TYPE "UDT_ZoneStructure"
VERSION : 0.1
   STRUCT
      SpeedZoneStart : DWord;
      SpeedZoneEnd : DWord;
      Zone : Word;
      Description : String[10];
      LastZone : Bool;
      StartPos : DWord;
      SpeedZone : Bool;
      NextZone : Int;
      PrevZone : Int;
      EndPos : DWord;
      AccumZone : Bool;
      ProductionZone : Bool;
      ProductionZoneSpacing : Word;
      MaxCarriers : Word;
      CarrierSpacing : Word;
      ClearToEnter : Bool;
      ClearOfStop : Bool;
      ClearZoneStart : Bool;
      ZoneFull : Bool;
      CarrierZnStatus : Array[0..60] of "UDT_ZoneCarrierStatus";
      CarrierZnStatusUnsorted : Array[0..60] of "UDT_ZoneCarrierStatus";
      InPositionTolerance : Word;
      NextCarrierClrHighSpeed : Word;
      DecelPositionOffset : Word;
      GapSpacingFault : Bool;
      GapFaultZnPosition : Int;
      GapFaultInZone : Int;
      FirstCarrierNumGapFlt : Int;
      SecondCarrierNumGapFlt : Int;
      FinePosStopZone : Bool;
      FineInPosTolerance : Word;
      FinePositionDecelOffset : Word;
      CoarseInPosTolerance : Word;
      CoarsePositionDecelOffset : Word;
      ZoneLength : Word;
      HMIZonePositionStatus : Array[1..20] of "UDT_HMIZonePositionStructure";
      HMIZonePositions : Array[1..20] of "UDT_HMIZonePositions";
      CarrierAtStop : Bool;
      CarrierNumAtStop : Word;
      StopControlFromEMS01 : "UDT_StopControlFromEMS01";
      ClearOfStopPos : DWord;
      StopStatusToEMS01 : "UDT_StopStatusToEMS01";
   END_STRUCT;
END_TYPE

TYPE "UDT_CarrierStructure"
VERSION : 0.1
   STRUCT
      SDC_IN : "UDT_SDC_IN";
      SDC_OUT : "UDT_SDC_OUT";
      ZoneFound : Word;
      Position : DWord;
      SpeedSelect : Word;
      MoveFWD : Bool;
      InProductionHold : Bool;
      Zone : Word;
      Area : String[2];
      AutoSpeedFast : Word;
      AutoSpeedSlow : Word;
      InPositionTolerance : Word;
      DecelSpeed : Word;
      DecelStartPos : DWord;
      ZonePosition : Word;
      CommFlt : Bool;
      CarrierPosition : DWord;
      CarrierNumber : Word;
      FaultsMasked : Bool;
      Faulted : Bool;
   END_STRUCT;
END_TYPE

TYPE "UDT_Zone"
VERSION : 0.1
   STRUCT
      ZONE : Array[1..60] of "UDT_ZoneStructure";
   END_STRUCT;
END_TYPE

TYPE "UDT_ZoneCarrierStatus"
VERSION : 0.1
   STRUCT
      CarrierNumber : Word;
      Position : DWord;
      RunningFWD : Bool;
   END_STRUCT;
END_TYPE

TYPE "UDT_OUT"
   STRUCT
      DecrementCarrierIndex : Bool;
      IncrementCarrierIndex : Bool;
      CarrierStatusIndex : Int;
      DecrementStatusIndex : Bool;
      IncrementStatusIndex : Bool;
      DriveStatusIndex : Int;
      DecrementZoneIndex : Bool;
      IncrementZoneIndex : Bool;
      ZoneStatusIndex : Int;
   END_STRUCT;
END_TYPE

TYPE "UDT_Carrier_Drive_Data"
   STRUCT
      CARRIER : Array[1..99] of "UDT_Drive_Data";
   END_STRUCT;
END_TYPE

TYPE "UDT_Drive_Data"
   STRUCT
      Drive_Control : Word;
      Drive_Status : Word;
   END_STRUCT;
END_TYPE

TYPE "UDT_Carrier_IO_HMI"
   STRUCT
      Carrier_Slot02_Inputs : Byte;
      Carrier_Slot03_Outputs : Byte;
      Carrier_Slot04_Inputs : Word;
      Carrier_Slot05_Outputs : Word;
   END_STRUCT;
END_TYPE

TYPE "UDT_IO_Data"
   STRUCT
      Slot2SafeInputs : Byte;
      Slot3SafeOutputs : Byte;
      Slot4StdInputs : Word;
      Slot5StdOutputs : Word;
   END_STRUCT;
END_TYPE

TYPE "UDT_Carrier_IO_Data"
   STRUCT
      CARRIER : Array[1..99] of "UDT_IO_Data";
   END_STRUCT;
END_TYPE

TYPE "UDT_Carrier_Status_HMI"
   STRUCT
      CarrierPosition : DWord;
      ActualSpeed : Word;
      RunningFWD : Bool;
      RunningREV : Bool;
      ProductionHoldPB_Status : Bool;
      CrashDetectStatus : Bool;
      AutoMode : Bool;
      ManualMode : Bool;
      DriveFwdCMD : Bool;
      DriveCmdSpeed : Word;
      NextCarrierNum : Word;
      NextStopPosition : DWord;
      Zone : Int;
      Area : String[2];
      CarrierFaultCode : Int;
      AtCmdPos : Bool;
      CommFlt : Bool;
      Faulted : Bool;
      CarrierStatusIndex : Int;
      DriveStatusIndex : Int;
      ZoneStatusIndex : Int;
      EncoderCommFault : Bool;
      DriveCommFault : Bool;
      HMICommFault : Bool;
      SetMaskCarrierFaultsPB : Bool;
      MaskCarrierFaultsLT : Bool;
      ResetMaskCarrierFaultsPB : Bool;
   END_STRUCT;
END_TYPE

TYPE "UDT_Zone_Status_HMI"
   STRUCT
      ZoneIndex : Int;
      ZoneType : String;
      NextZoneNumber : Int;
      ZoneStartPosition : DWord;
      ZoneEndPosition : DWord;
      ZoneFull : Bool;
      SpeedZone : Bool;
      SpeedZoneStartPos : DWord;
      SpeedZoneEndPos : DWord;
      AccumZoneSpacing : Word;
      ProductionZoneSpacing : Word;
      CarrierZoneStatus : Array[0..60] of "UDT_ZoneCarrierStatus";
   END_STRUCT;
END_TYPE

TYPE "UDT_StopStatusToEMS01"
   STRUCT
      StopOpen : Bool;
      StopClosed : Bool;
      CarrierAtStop : Bool;
      CarrierReleasingFromStop : Bool;
   END_STRUCT;
END_TYPE

TYPE "UDT_StopControlFromEMS01"
   STRUCT
      ClearToOpen : Bool;
      ClearToReleaseCarrier : Bool;
   END_STRUCT;
END_TYPE

TYPE "UDT_G120D_STW1_CONTROL"
VERSION : 0.1
   STRUCT
      Bit_08_JOG_R : Bool;   // 1=tippen rechtsseitig EIN/ 0= AUS / 1=jogging on right-hand side ON/ 0= OFF
      Bit_09_JOG_L : Bool;   // 1=tippen linksseitig EIN/ 0= AUS / 1=jogging on left-hand side ON/ 0= OFF
      Bit_10_CONTR_PLC : Bool;   // 1=Bedienung über PLC erforderlich/ 0=keine Bedienung über PLC erforderlich / 1=control by PLC required/ 0=no control by PLC required
      Bit_11_REVERSE : Bool;   // 1=Umkehrung des Sollwerts/ 0=keine Umkehrung / 1=inversion of setpoint/ 0=no inversion of setpoint
      Bit_12_BRAKE_Release : Bool;   // 1= Löse Bremse / 1= Release Break / 1= Manual Brake Release
      Bit_13_DDS : Bool;   // 1=DDS1 FU Datenset / 0=DDS0 FU Datenset / 1=DDS1 FU Dataset / 0=DDS0 FU Dataset
      Bit_14_DO0 : Bool;   // 1=Digitaler Ausgang aktiv/ 0=Digitaler Ausgang nicht aktiv / 1=Digital Output activ/ 0=Digital Output not activ
      Bit_15_DO1 : Bool;   // 1=Digitaler Ausgang aktiv/ 0=Digitaler Ausgang nicht aktiv / 1=Digital Output activ/ 0=Digital Output not activ
      Bit_00_ON : Bool;   // 1=EIN/ 0=AUS / 1=ON/ 0=OFF2
      Bit_01_AUS2_INH : Bool;   // 1=Betriebsvoraussetzung/ 0=AUS2 - Pulsverzögerer, Spannung auf einmal aus / 1=operation condition/ 0=AUS2 - pulse inhibitor, voltage off at once
      Bit_02_AUS3_STOP : Bool;   // 1=Betriebsvoraussetzung / 0=AUS3 - schneller Halt / 1=operation condition / 0=AUS3 - fast stop
      Bit_03_EN : Bool;   // 1=Freigabe Betrieb/ 0=deaktiviere Betrieb / 1=enable operation/ 0=disable operation
      Bit_04_EN_RAMP : Bool;   // 1=1=Betriebsvoraussetzung / 0=deaktiviere Funktionsrampengenerator / 1=operation condition / 0=disable ramp function generator
      Bit_05_START_RAMP : Bool;   // 1=Aktiviere Rampenfunktion / 0=deaktivere RFG / 1=enable ramp function generator / 0=stoppen RFG
      Bit_06_SETPOINT : Bool;   // 1=Freigabe Sollwert/ 0=deaktiviere Sollwert / 1=enable setpoint/ 0=disable setpoint
      Bit_07_RESET : Bool;   // 1=Störung quittieren / 0= irrelevant / 1=Reset fault / 0= irrelevant
   END_STRUCT;
END_TYPE

TYPE "UDT_G120D_ZSW1_STATUS"
VERSION : 0.1
   STRUCT
      Bit_08_NO_DEVIATION : Bool;   // 1=keine Abweichung des Sollwerts / 0=Abweichung / 1=no deviation current-setpoint / 0=deviation / Setpoint / actual value deviation within the tolerance range.
      Bit_09_CONTR_PLC : Bool;   // 1=Kontrolle über PLC erforderlich/ 0=keine Kontrolle erforderlich / 1=control by PLC required/ 0=no control by PLC required / The automation system is requested to ac-cept the inverter control.
      Bit_10_F_MAX : Bool;   // 1=fmax erreicht/ 0= unter fmax / 1=fmax reached/ 0= below fmax / Speed is greater than or equal to the corre-sponding maximum speed.
      Bit_11_LIMIT_REACHED : Bool;   // 1=keine Warnung/ 0=Warnung: Motor an Spannungsgrenze / 1=no warning/ 0=warning:Motor at limit of current / Comparison value for current or torque has been reached or exceeded.
      Bit_12_BRAKE_OPEN : Bool;   // 1= / 0=Haltebremse / motor Brake is open
      Bit_13_NO_OVERTEMP : Bool;   // 1= / 0=Motorüberlast / Drive Overtemperature
      Bit_14_CW_CCW : Bool;   // 1=Rechtslauf/ 0=Linkslauf / On for drive runnin clockwise/off counterclockwise
      Bit_15_OVERL : Bool;   // 1= /0= Konvertierer Überlast / 1= /0= Konverter overload / 0 = Alarm, in-verter thermal overload/on CDS display
      Bit_00_READY_RUN : Bool;   // 1=bereit zum betreiben/ 0= nicht bereit / 1=ready to run/ 0= not ready to run / Power supply switched on; electronics initial-ized; pulses locked.
      Bit_01_READY_ON : Bool;   // 1=bereit zum einschalten/ 0= nicht bereit / 1=ready to switch on/ 0= not ready to switch on / Motor is switched on (ON/OFF1 = 1), no fault is active. With the command "Enable opera-tion" (STW1.3), the inverter switches on the motor.
      Bit_02_ENABLE : Bool;   // 1=Freigabe Bedienung / 0=deaktiviere Bedienung / 1=operation enabled / 0=operation disabled / Motor follows setpoint. See control word 1, bit 3.
      Bit_03_FAULT : Bool;   // 1=Störung / 0=keine Störung / 1=fault / 0=no fault / The inverter has a fault. Acknowledge fault using STW1.7
      Bit_04_OFF2 : Bool;   // 1=kein AUS2 / 0=AUS2 Befehl ist vorhanden / 1=no AUS2 / 0=AUS2 command is present / OFF2 Coast down to standstill is not active.
      Bit_05_OFF3 : Bool;   // 1=kein AUS3 / 0=AUS3 Befehl ist vorhanden / 1=no AUS3 / 0=AUS3 command is present / OFF3 Quick stop is not active.
      Bit_06_LOCK_OUT : Bool;   // 1=sperre Ausschaltung / 0=keine Sperrung / 1=closing lock-out / 0=no closing lock-out / It is only possible to switch on the motor after an OFF1 followed by ON.
      Bit_07_WARN : Bool;   // 1=Warnung / 0= keine Warnung / 1=Warning / 0= no warning
   END_STRUCT;
END_TYPE

TYPE "UDT_G120D_ERRORS"
VERSION : 0.1
   STRUCT
      F_X33_F1 : Bool;   // Fehler Überstrom
      F_X34_F2 : Bool;   // Fehler Überspannung
      F_X35_F3 : Bool;   // Fehler Unterspannung
      F_X36_F4 : Bool;   // Fehler Inverter Übertemperatur
      F_X37_F41 : Bool;   // Fehler Motordatenerkennung
      F_X38_F52 : Bool;   // Fehler Leistungsteil
      F_X39_F62 : Bool;   // Fehler MMC Daten sind fehlerhaft
      F_X40_F70 : Bool;   // Fehler PLC Sollposition
      F_X41_F71 : Bool;   // Fehler USS Sollposition, Überwachung
      F_X42_F72 : Bool;   // Fehler USS Sollposition, USS Master
      F_X43_F90 : Bool;   // Fehler Gebersignal
      F_X44_F395 : Bool;   // Fehler CU/PM wechsel
      bit_14 : Bool;   // Reserve
      bit_15 : Bool;   // Reserve
      bit_16 : Bool;   // Reserve
      bit_17 : Bool;   // Reserve
   END_STRUCT;
END_TYPE

TYPE "UDT_SDC_EMS_FLAGS"
VERSION : 0.1
   STRUCT
      PRESENT : Bool;   // EMS vorhanden
      IN_HW : Bool;   // EMS in HardwareConfiguration
      ACTIV : Bool;   // EMS activiert
      ENABLE : Bool;   // EMS enable
      COMM_FAULT : Bool;   // EMS communicationsfehler
      FAULTY : Bool;   // EMS fehlerhaft
      SIMULATION : Bool;   // EMS simualtion
      Spare_0_7 : Bool;   // Spare
      Spare_1_0 : Bool;   // Spare
      Spare_1_1 : Bool;   // Spare
      Spare_1_2 : Bool;   // Spare
      Spare_1_3 : Bool;   // Spare
      Spare_1_4 : Bool;   // Spare
      Spare_1_5 : Bool;   // Spare
      Spare_1_6 : Bool;   // Spare
      Spare_1_7 : Bool;   // Spare
   END_STRUCT;
END_TYPE

TYPE "UDT_SDC_TS_PARAMETER"
VERSION : 0.1
   STRUCT
      ALLG : "UDT_SDC_TS_PAR_ALLG";   // allgemeine Sections Parameter
      PROFIL : Array[1..10] of "UDT_SDC_TS_PAR_PROFIL";   // Profilbezogene Sections Parameter
   END_STRUCT;
END_TYPE

TYPE "UDT_SDC_TS_PAR_PROFIL"
VERSION : 0.1
   STRUCT
      Hoist_Pos_start : Int;   // Start of hoist positioning; offset from start pos.(mm)
      Height : Int := 2651;   // Setpoint: hoist position (mm)
      Hoist_speed : Int := 2000;   // Setpoint: hoist speed (mm/min)
      Hoist_offset_1 : Int;   // set value: hoist offset (mm)
      Hoist_offset_2 : Int;   // set value: hoist offset (mm)
      Hoist_offset_3 : Int;   // set value: hoist offset (mm)
      Hoist_offset_4 : Int;   // set value: hoist offset (mm)
      Hoist_Start_offset_1 : Int;   // Start der Hubbewegung zu offset 1, Offset von Startpos. (mm)
      Hoist_Start_offset_2 : Int;   // Start der Hubbewegung zu offset 1, Offset von Startpos. (mm)
      Hoist_Start_offset_3 : Int;   // Start der Hubbewegung zu offset 1, Offset von Startpos. (mm)
      Hoist_Start_offset_4 : Int;   // Start der Hubbewegung zu offset 1, Offset von Startpos. (mm)
   END_STRUCT;
END_TYPE

TYPE "UDT_SDC_TS_PAR_ALLG"
VERSION : 0.1
   STRUCT
      SEK_NEXT_1 : Int;   // Sektion next 1
      SEK_NEXT_2 : Int;   // Sektion next 2
      Spare : Array[4..5] of Byte;   // Spare
      POS : "UDT_SDC_TS_PAR_POS";   // Pos Parameter
      FLAGS : Struct
         DIST_VAL : Array[0..15] of Bool;   // Abstandswerte
         one_profile : Bool;   // Reserved for: only one profile
         BLIND : Bool;   // Reserved for: Blind travel without position values
         NO_DIST_CONT : Bool;   // without distance control (no slow speed, ...)
         SYNCH_AREA : Bool;   // synchronous conveyor area
         bit24 : Bool;   // spare
         bit25 : Bool;   // spare
         bit26 : Bool;   // spare
         bit27 : Bool;   // spare
         EN_HOIST : Bool;   // Hoist/tilt enable
         D_RESET_AFTER : Bool;   // Antrieb belegt nach Reset vorhanden
         D_PULK : Bool;   // Antriebs PULK
         bit33 : Bool;   // spare
         bit34 : Bool;   // spare
         bit35 : Bool;   // spare
         bit36 : Bool;   // spare
         Deutronic_ON : Bool;   // Reserved for: DEUTRONIC CHARGE COMPUTER ON
      END_STRUCT;
      Stop_Position : Int;   // Stopp position, offset from start pos.(mm)
      Drive_speed_1 : DInt;   // set value: drive speed (mm/min)
      Drive_speed_2 : DInt;   // set value: drive speed (mm/min)
   END_STRUCT;
   // FLAGS.DIST_VAL[0] := true;
END_TYPE

TYPE "UDT_SDC_TS_PAR_POS"
VERSION : 0.1
   STRUCT
      Start_1 : DInt := 0;   // mm
      End_1 : DInt := 0;   // mm
      Start_2 : DInt;   // Reserve
      End_2 : DInt;   // Reserve
      Actionpoint_1 : Int;   // Fahrantrieb Aktionspunkt 1
      Actionpoint_2 : Int;   // Fahrantrieb Aktionspunkt 2
   END_STRUCT;
END_TYPE

TYPE "UDT_EMS_IF_Q"
VERSION : 0.1
   STRUCT
      STAT : "UDT_EMS_IF_Q_STAT";   // Statusbit`s / Stausbit`s
      ERROR : Int;   // Störnummer / Error number
      D_POS : DInt;   // Fahrantrieb Position in mm / Drive position in mm
      H_POS : Int;   // Hubantrieb Position in mm / Hoist position in mm
      SPARE_POS : Int;
      VFC : "UDT_EMS_IF_Q_VFC";   // Prozesswerte FU`s / Processdata VFC
      IQ : "UDT_EMS_IF_Q_IQ";   // Ein-Ausgänge / In-Outputs
      ER_WORD_No : Int;   // Zähler Störnummern / Counter error words
      ER_WORD : Word;   // Datenwort Störnummern / Dataword error words
      FB_DBNo : Int;   // Rückmeldung DB Nummer Datentransfer / Feedback DB No. data transfer
      FB_DBBNo : Int;   // Rückmeldung DBB Nummer Datentransfer / Feedback DBB No. data transfer
   END_STRUCT;
END_TYPE

TYPE "UDT_SDC_EMS"
VERSION : 0.1
   STRUCT
      IF_I_EMS : "UDT_EMS_IF_Q";   // Inputs from EMS
      IF_Q_EMS : "UDT_EMS_IF_I";   // Outputs to EMS
      TS_PAR : Struct   // Section parameters
         ALLG : "UDT_SDC_TS_PAR_ALLG";   // Section parameters allg
         PROFIL : "UDT_SDC_TS_PAR_PROFIL";   // Section parameters Profil
      END_STRUCT;
      TS_STAT : "UDT_SDC_EMS_TS_STAT";   // EMS Sektion Stat Daten
      TS_COM : "UDT_SDC_EMS_TS_COM";   // EMS Sektion Com Daten
      FKT : "UDT_SDC_EMS_FKT_BITs";   // EMS Funktionen
      FKT_RESET : "UDT_SDC_EMS_FKT_BITs";   // EMS Funktionen reset
      FLAGS : "UDT_SDC_EMS_FLAGS";   // EMS Fahnen
      FKT_INFO_REP_1 : Int;   // EMS Funktionen Info Repair 1
      FKT_INFO_REP_2 : Int;   // EMS Funktionen Info Repair 2
      PROFIL : Int;   // Profile Number
      CYCLE_COUNTER : Int;   // Zykluszähler
      PRECEDING_EMS : Int;   // preciding EMS
      DISTANCE : DInt;   // Abstand zum vorangehenden EMS
      ABS_POS : DInt;   // absolute Positon
      NewSektion : Bool;   // New Sektion
      BcOk : Bool;   // Barcode ist OK
      SekOk : Bool;   // Sektion is OK
      Spare_0_3 : Bool;   // Spare
      Spare_0_4 : Bool;   // Spare
      Spare_0_5 : Bool;   // Spare
      Spare_0_6 : Bool;   // Spare
      Spare_0_7 : Bool;   // Spare
      Send_EMS_PAR_Act : Bool;   // Sende EMS Parameter aktiv
      Send_EMS_PAR_End : Bool;   // Sende EMS Parameter ende
      Send_EMS_LEAPS_Act : Bool;   // Sende EMS Sprünge aktiv
      Send_EMS_LEAPS_End : Bool;   // Sende EMS Sprünge ende
      H_C_Pos : Array[0..4] of Bool;   // Hub Kommando positionierung / Offset 1 / ,...
      Spare246 : Array[246..249] of Byte;   // Spare
      ER : "UDT_EMS_IF_I_SDC_ERRORS";
      WA_DIST : Bool;   // Warning Distance
      WA_COLL : Bool;   // Warning Collision Sensor activ
      WA_DIST_SAFETY : Bool;   // Warning Distance safety
      WA_Spare_2_3 : Bool;   // Warning Spare 2.3
      WA_Spare_2_4 : Bool;   // Warning Spare 2.4
      WA_Spare_2_5 : Bool;   // Warning Spare 2.5
      WA_Spare_2_6 : Bool;   // Warning Spare 2.6
      WA_Spare_2_7 : Bool;   // Warning Spare 2.7
      WA_Spare_3 : Byte;   // Warning Spare 3
      Spare254 : Array[254..257] of Byte;   // Spare
      VersNo : Array[0..1] of Byte;
   END_STRUCT;
END_TYPE

TYPE "UDT_SDC_EMS_TS_STAT"
VERSION : 0.1
   STRUCT
      VAL : "UDT_SDC_TS_IF_STATUS_VAL";
      BIT : "UDT_SDC_TS_IF_STATUS_BIT";
      SORTE : Array[1..4] of Char;   // Karossentyp
      FKT : "UDT_SDC_EMS_FKT_BITs";
      SPARE : Word;
   END_STRUCT;
END_TYPE

TYPE "UDT_SDC_EMS_TS_COM"
VERSION : 0.1
   STRUCT
      VAL : "UDT_SDC_TS_IF_COMMAND_VAL";
      BIT : "UDT_SDC_TS_IF_COMMAND_BIT";
      FKT_SET : "UDT_SDC_EMS_FKT_BITs";
      FKT_RESET : "UDT_SDC_EMS_FKT_BITs";
   END_STRUCT;
END_TYPE

TYPE "UDT_EMS_IF_Q_STAT"
VERSION : 0.1
   STRUCT
      LIFE_BIT : Bool;   // Lebensbit / Heartbeat
      ER_SUM : Bool;   // Sammelfehler / Summaryerror
      IR_MAN : Bool;   // EMS in Handbetrieb / EMS in manual mode (IR)
      ER_RESET : Bool;   // Störung quittieren / Error reset (IR)
      HOIST_CLEAR : Bool;   // Hub über/in Sollpos und Bereit ohne Störung / Hoist above position and no error
      POS_START_X : Bool;   // Fahrantrieb positioniert / Drive positioning started
      ALWAYS_ONE : Bool;   // immer "1" / Always "1"
      H_DISABLED : Bool;   // Hub gesperrt / Hoist disabled
      D_FWD : Bool;   // Fahrantrieb fährt vorwärts / Drive moves forwards
      D_RWD : Bool;   // Fahrantrieb fährt rückwärts / Drive moves reward
      bit12 : Bool;   // Reserve / spare
      D_IN_POS : Bool;   // Fahrantrieb in Position / Drive in Position
      H_UP : Bool;   // Hub hebt / Hoist raises
      H_DOWN : Bool;   // Hub senkt / Hoist lowers
      H_IN_POS : Bool;   // Hub in Position / Hoist in position
      H_IN_TOPPOS : Bool;   // Hub in oberster Position / Hoist in top position
      bit2_0 : Bool;   // Schwenkantrieb fährt + / Tilt moves clockwise
      bit2_1 : Bool;   // Schwenkantrieb fährt - / Tilt moves counterclockwise
      bit2_2 : Bool;   // Hub in oberster Position / Tilt in position
      bit2_3 : Bool;   // Hub in Grundstellung / Tilt in home position
      IN_BOTPOS : Bool;   // Hub in unterster Position / Hoist In bottom Position (min) (with Tiltposition)
      bit2_5 : Bool;   // Reserve / spare
      bit2_6 : Bool;   // Reserve / spare
      bit2_7 : Bool;   // Reserve / spare
      MESS_ACT : Bool;   // Störnummer ist eine Meldung / Error No is a Message
      MESS_POS : Bool;   // Reserve / spare
      bit3_2 : Bool;   // Reserve / spare
      bit3_3 : Bool;   // Reserve / spare
      bit3_4 : Bool;   // Reserve / spare
      bit3_5 : Bool;   // Reserve / spare
      bit3_6 : Bool;   // Reserve / spare
      DATA_TRANS : Bool;   // Datentransfer ist aktiv / Data Transfer aktiv
   END_STRUCT;
END_TYPE

TYPE "UDT_EMS_IF_I_CONTR"
VERSION : 0.1
   STRUCT
      LIFE_BIT : Bool;   // Lebensbit / Heartbeat
      ER_SDC : Bool;   // Sammelfehler / Summaryerror
      H_EMERG : Bool;   // Hubantrieb Notbetrieb / Hoist Emergency mode
      Spare_0_3 : Bool;   // Schwenkantrieb Notbetrieb / Tilt Emergency mode
      LAMP_TEST : Bool;   // Lampentest / Lamp Test
      VAC_CLEAN : Bool;   // EMS mit Staubsauger / EMS with vac cleaner
      SYNCH : Bool;   // Synchronbetrieb / Control distance, synchronous area
      DATA_TRANS : Bool;   // Datentransfer ist aktiv / Data Transfer aktiv
      ER_RESET : Bool;   // Störung quittieren / Error reset
      AUTO : Bool;   // 1 = Automatikbetrieb / Automatic mode in section
      MAN : Bool;   // 1 = Handbetrieb / Manual mode in section
      D_C_BREAK : Bool;   // Fahrantrieb Befehl Bremse lüften / DRIVE Command release Break
      H_C_BREAK : Bool;   // Hubantrieb Befehl Bremse lüften / HOIST Command release Break
      D_EMERG_FC : Bool;   // Fahrantrieb Notbetrieb 1 Motor / DRIVE Emergency mode Frequencyconverter 1 Motor
      INC_TOL_POS : Bool;   // Schwenkantrieb Notbetrieb 1 Motor / TILT Emergency mode Frequencyconverter 1 Motor
      E_STOP : Bool;   // "1"Not-Halt / Emergency stop from Interface
      D_C_FWD : Bool;   // Fahrantrieb Befehl vorwärts / DRIVE Command forward
      D_C_RWD : Bool;   // Fahrantrieb Befehl rückwärts / DRIVE Command reward
      D_C_BSP : Bool;   // Fahrantrieb Befehl weiter fahren / DRIVE Command bridge stop position
      Spare_2_3 : Bool;   // Reserve / spare
      IR_noEMSnumber : Bool;   // Schwenkantrieb Befehl + / TILT Command clockwise
      IR_noLogin : Bool;   // Schwenkantrieb Befehl - / TILT Command counterclockwise
      BYP_scalance_PN_error : Bool;   // Schwenkantrieb Befehl positionieren / TILT Command positioning
      Spare_2_7 : Bool;   // Schwenkantrieb Befehl fahren in Grundstellung / TILT Command to home position, high priority
      H_C_UP : Bool;   // Hubantrieb Befehl heben / HOIST Command raise without positioning
      H_C_DOWN : Bool;   // Hubantrieb Befehl senken / HOIST Command lower without positioning
      H_C_POS : Bool;   // Hubantrieb Befehl positionieren / HOIST Command hoist positioning
      H_C_TOP : Bool;   // Hubantrieb Befehl fahren in oberste Position / HOIST Command Raise to top position, high priority
      H_EN : Bool;   // Hub-Schwenkfreigabe / HOIST-TILT enable
      H_BYP_ROPE : Bool;   // Überbrücken Seilkontrolle / Bypass monitoring of rope
      Spare_3_6 : Bool;   // Reserve / spare
      H_BYP_REF_INI : Bool;   // Überbrücken Kontrolle Referenzinitiator (nicht safety) / No monitoring of reference initiator (non safety)
   END_STRUCT;
END_TYPE

TYPE "UDT_SDC_TS_IF_COMMAND_BIT"
AUTHOR : SIEMENS
FAMILY : FT
NAME : SDC_BIT
VERSION : 2.0
   STRUCT
      ER_RESET : Bool;   // Error Reset
      AUTO : Bool;   // 1 = Automatik in Sektion
      MAN : Bool;   // 1 = Handbetrieb in Sektion
      Spare_0_3 : Bool;   // Reserve
      Spare_0_4 : Bool;   // Reserve
      E_STOP : Bool;   // "1" -> NotAus von Interface (system PLC)
      Spare_0_6 : Bool;   // Reserve
      Spare_0_7 : Bool;   // Reserve
      D_C_FWD : Bool;   // Fahrantrieb Kommando vorwärts
      D_C_RWD : Bool;   // Fahrantrieb Kommando rückwärts
      D_C_BSP : Bool;   // Fahrantrieb Kommando Überbrückung Stopp-Position
      D_C_V1 : Bool;   // Fahrantrieb Kommando Geschwindigkeit 1
      D_C_V2 : Bool;   // Fahrantrieb Kommando Geschwindigkeit 2
      D_C_V_VAR : Bool;   // Fahrantrieb Kommando variabler Geschwindigkeit
      D_C_BEFOR_POS : Bool;   // Fahrantrieb Kommando Freigabe vor Stop-Position
      D_C_AFTER_POS : Bool;   // Fahrantrieb Kommando Freigabe nach Stop-Position
      H_C_RAISE : Bool;   // Hubantrieb Kommando aufwärts
      H_C_LOWER : Bool;   // Hubantrieb Kommando abwärts
      H_C_POS : Bool;   // Hubantrieb Kommando Positionieren
      H_C_POS1 : Bool;   // Hubantrieb Kommando Offset 1
      H_C_POS2 : Bool;   // Hubantrieb Kommando Offset 2
      H_C_POS3 : Bool;   // Hubantrieb Kommando Offset 3
      H_C_POS4 : Bool;   // Hubantrieb Kommando Offset 4
      H_C_TOP : Bool;   // Hubantrieb Kommando nach Top Position, hohe Priorität
      H_BYP_ROPE : Bool;   // Hubantrieb Überbrücken Seilkontrolle
      Spare_3_1 : Bool;   // Reserve
      H_BYP_REF_INI : Bool;   // Hubantrieb Überbrücken Kontrolle Referenzinitiator (nicht safety)
      H_C_SLOW : Bool;   // Hubantrieb Kommando globaler Parameter langsam
      D_BYP_DIST_CONTR : Bool;   // Fahrantrieb Überbrücke Distanzkontrolle
      Spare_3_5 : Bool;   // Reserve
      Spare_3_6 : Bool;   // Reserve
      SET_PROF : Bool;   // setze Profile
   END_STRUCT;
END_TYPE

TYPE "UDT_SDC_TS_IF_COMMAND_VAL"
AUTHOR : SIEMENS
FAMILY : FT
NAME : SDC_VAL
VERSION : 1.6
   STRUCT
      PROFIL : Int;   // Profile
      D_SETSPEED : DInt;   // set value: drive speed (mm/min)
      D_POS_OFFS : Int;   // Antriebsposition offset
      H_POS_OFFS : Int;
   END_STRUCT;
END_TYPE

TYPE "UDT_SDC_TS_IF_STATUS_BIT"
AUTHOR : SIEMENS
FAMILY : FT
NAME : SDC_BIT
VERSION : 1.6
   STRUCT
      PRESENT : Bool;   // EMS vorhanden
      ERROR : Bool;   // Sammelstörung
      MAN_IR : Bool;   // EMS in Handbetrieb (Fernsteuerung)
      MORE_EMS_PRESENT : Bool;   // Mehr als 1 EMS in Sektion vorhanden
      ER_COMMAND : Bool;   // Fehlerhafte Befehle von System PLC
      W_DIST : Bool;   // Warnung Distanckontrolle ist aktiv
      Spare_0_6 : Bool;   // Warnung Auffahrsensor ist aktiv Reserve
      MESS_ACT : Bool;   // Störnummer ist eine Meldung / Error No is a Message
      D_MOVING : Bool;   // Fahrantrieb ist ein
      D_NOT_MOVING : Bool;   // Fahrantrieb ist aus
      H_MOVING : Bool;   // Hubantrieb ist ein
      H_NOT_MOVING : Bool;   // Hubantrieb ist aus
      X_MOVING : Bool;   // Reserve Antrieb ein
      X_NOT_MOVING : Bool;   // Reserve Antrieb aus
      D_IN_POS : Bool;   // Fahrantrieb in Position
      Spare_2_1 : Bool;   // Reserve
      D_BEFOR_POS : Bool;   // Fahrantrieb vor Stopposition
      D_AFTER_POS : Bool;   // Fahrantrieb nach Stopposition
      D_GR_AP1 : Bool;   // Fahrantrieb Barcodeposition größer Aktionspunkt 1
      D_SM_AP1 : Bool;   // Fahrantrieb Barcodeposition kleiner Aktionspunkt 1
      D_GR_AP2 : Bool;   // Fahrantrieb Barcodeposition größer Aktionspunkt 2
      D_SM_AP2 : Bool;   // Fahrantrieb Barcodeposition kleiner Aktionspunkt 2
      H_IN_POS : Bool;   // Hubantrieb in Position (hoist drive)
      H_IN_TOPPOS : Bool;   // Hubantrieb in top pos.(limit)
      H_IN_POS1 : Bool;   // Hubantrieb in Position (hoist drive) Offset 1
      H_IN_POS2 : Bool;   // Hubantrieb in Position (hoist drive) Offset 2
      H_IN_POS3 : Bool;   // Hubantrieb in Position (hoist drive) Offset 3
      H_IN_POS4 : Bool;   // Hubantrieb in Position (hoist drive) Offset 4
      H_GR_POS : Bool;   // Hubposition größer Sollposition ohne Offset
      H_SM_POS : Bool;   // Hubposition kleiner Sollposition ohne Offset
      H_GR_POS1 : Bool;   // Hubposition größer Sollposition + Offset 1
      H_SM_POS1 : Bool;   // Hubposition kleiner Sollposition + Offset 1
      H_GR_POS2 : Bool;   // Hubposition größer Sollposition + Offset 2
      H_SM_POS2 : Bool;   // Hubposition kleiner Sollposition + Offset 2
      H_GR_POS3 : Bool;   // Hubposition größer Sollposition + Offset 3
      H_SM_POS3 : Bool;   // Hubposition kleiner Sollposition + Offset 3
      H_GR_POS4 : Bool;   // Hubposition größer Sollposition + Offset 4
      H_SM_POS4 : Bool;   // Hubposition kleiner Sollposition + Offset 4
      H_BOTTOM_POS : Bool;   // Hub (mit Neigung) in unterer Position
      H_DISABLED : Bool;   // Hub ist verriegelt, keine Freigabe
      H_CLEAR : Bool;   // Hub über/in Sollpos und bereit ohne Störung
      D_MOVING_FWD : Bool;   // Fahrantrieb Bewegung vorwärts
      D_MOVING_RWD : Bool;   // Fahrantrieb Bewegung rückwärts
      D_RESET_AFTER : Bool;   // Fahrantrieb Bewegung Belegt Reset ohne Present
      D_PULK : Bool;   // Fahrantrieb Sektion in PULKbetrieb
      D_NO_POS : Bool;   // Fahrantrieb keine Stopposition Sektion
      Spare_7_6 : Bool;
      Spare_7_7 : Bool;
   END_STRUCT;
END_TYPE

TYPE "UDT_SDC_TS_IF_STATUS_VAL"
AUTHOR : SIEMENS
FAMILY : FT
NAME : SDC_VAL
VERSION : 1.6
   STRUCT
      EMS_ID : Int;   // EMS ID Nummer
      PROFIL : Int;   // Profile
      DRIVE_POS : DInt;   // Antriebsposition in mm
      HOIST_POS : Int;   // Höhe in mm
      ERROR : Int;   // Error-Nummer
      DRIVE_POS_PERC : Int;   // Position [% of Start End Section]
      SEK : Int;   // Sektion
   END_STRUCT;
END_TYPE

TYPE "UDT_SDC_EMS_FKT_BITs"
VERSION : 0.1
   STRUCT
      EMS_TO_REPAIR_1 : Bool;   // EMS zur Reperatur 1
      EMS_TO_REPAIR_2 : Bool;   // EMS zur Reperatur 2
      EMERG_HOIST : Bool;   // EMS Emergancy without Hoist
      Reserve_03 : Bool;   // EMS Emergancy without Tilt
      EMERG_DRIVE_FC : Bool;   // EMS Drive Emergency mode Frequencyconverter 1 Motor
      Reserve_05 : Bool;   // EMS Tilt Emergency mode Frequencyconverter 1 Motor
      LAMP_TEST : Bool;   // EMS Lamp Test
      VAC_CLEAN : Bool;   // EMS VAC Reiniger
      PE_TEST : Bool;   // EMS PE Test NIO
      KOHLE_TEST : Bool;   // EMS KOHLE Test NIO
      KOM_TEST : Bool;   // Reserve
      Reserve_11 : Bool;   // Reserve
      Reserve_12 : Bool;   // Reserve
      Reserve_13 : Bool;   // Reserve
      Reserve_14 : Bool;   // Reserve
      Reserve_15 : Bool;   // Reserve
   END_STRUCT;
END_TYPE

TYPE "UDT_EMS_IF_I_SDC_ERRORS"
VERSION : 0.1
   STRUCT
      _901_ER_SUM : Bool;   // Error SDC + EMS Summary
      _902_ER_SUM_SDC : Bool;   // Error SDC Summary
      _903_ER_BC_JUMP : Bool;   // Error SDC Barcode Jump
      _904_ER_NO_SEK : Bool;   // Error SDC no Section found
      _905_ER_COMMAND : Bool;   // Error SDC worng Commands from Main Plc
      _906_ER_BC_LIM : Bool;   // Error SDC Barcode LIMIT
      _907_ER_EMS_ID : Bool;   // Error SDC wrong EMS Number
      _908_ER_SEK_NR : Bool;   // Error SDC wrong Sektion Number
      _909_ER_LIFE : Bool;   // Error SDC Lifebeat to EMS
      _910_ER_BUS : Bool;   // Error SDC no Buscommunication to EMS device
      _911 : Bool;   // spare
      _912 : Bool;   // spare
      _913 : Bool;   // spare
      _914 : Bool;   // spare
      _915 : Bool;   // spare
      _916 : Bool;   // spare
   END_STRUCT;
END_TYPE

TYPE "UDT_SDC_ERROR_STAT"
VERSION : 0.1
   STRUCT
      EMS_TS_STAT_VAL : "UDT_SDC_TS_IF_STATUS_VAL";
      ER : "UDT_EMS_IF_I_SDC_ERRORS";
      Spare : Int;   // spare
      ER_DATE : Date_And_Time;   // Fehler Zeit
   END_STRUCT;
END_TYPE

// folder: UDT_AB_Interlocks

TYPE "UDT_AB_Interlocks_Carrier"
VERSION : 0.1
   STRUCT
      Carrier_IN : "UDT_AB_Interlocks_Carrier_In";
      Carrier_OUT : "UDT_AB_Interlocks_Carrier_Out";
   END_STRUCT;
END_TYPE

TYPE "UDT_AB_Interlocks_SDC_In"
VERSION : 0.1
   STRUCT
      EMS01_MasterPowerOn : Bool;
      EMS01_Fault_Reset_PB : Bool;
      EMS01R1_MasterPowerOn : Bool;
      EMS01R1_Fault_Reset_PB : Bool;
      EMS01R2_MasterPowerOn : Bool;
      EMS01R2_Fault_Reset_PB : Bool;
      EMS01R3_MasterPowerOn : Bool;
      EMS01R3_Fault_Reset_PB : Bool;
      EMS01R4_MasterPowerOn : Bool;
      EMS01R4_Fault_Reset_PB : Bool;
      EMS_Stop_26_Set_To_Release : Bool;
      Spare_11 : Bool;
      Spare_12 : Bool;
      Spare_13 : Bool;
      Spare_14 : Bool;
      Heartbeat : Bool;
      SpareWord2 : Word;
      SpareWord3 : Word;
      CarrierSpeedRef : Word;
      ProductionSpeedRef : Word;
   END_STRUCT;
END_TYPE

TYPE "UDT_AB_Interlocks_CarrierStatus_Out"
VERSION : 0.1
   STRUCT
      Spare0 : Bool;
      DriveTripped : Bool;
      Spare2 : Bool;
      PositioningComplete : Bool;
      RunStopPressed : Bool;
      Moving : Bool;
      Faulted : Bool;
      InAuto : Bool;
      Spare8 : Bool;
      Spare9 : Bool;
      Spare10 : Bool;
      Spare11 : Bool;
      Spare12 : Bool;
      Spare13 : Bool;
      Spare14 : Bool;
      Spare15 : Bool;
   END_STRUCT;
END_TYPE

TYPE "UDT_AB_Interlocks_Carrier_Out"
VERSION : 0.1
   STRUCT
      Status : "UDT_AB_Interlocks_CarrierStatus_Out";
      Fault : Word;
      Position : DWord;
      Zone : Word;
   END_STRUCT;
END_TYPE

TYPE "UDT_AB_Interlocks_Carrier_In"
VERSION : 0.1
   STRUCT
      CarrierDelete : Bool;
   END_STRUCT;
END_TYPE

TYPE "UDT_AB_Interlocks"